REGION Network 2
   RUNG wire#powerrail
      "DB204"(IN0 := "4#配料皮带备妥", IN1 := "干矿提升皮带运行", IN2 :=, IN3 :=, IN4 := "4#配料皮带运行", IN5 :=, OUT6 := "4#配料皮带启动")
      "DB205"(IN0 := "5#配料皮带备妥", IN1 := "干矿提升皮带运行", IN2 :=, IN3 :=, IN4 := "5#配料皮带运行", IN5 :=, OUT6 := "5#配料皮带启动")
      "DB206"(IN0 := "6#配料皮带备妥", IN1 := "干矿提升皮带运行", IN2 :=, IN3 :=, IN4 := "6#配料皮带运行", IN5 :=, OUT6 := "6#配料皮带启动")
   END_RUNG
   // the same network as SCL:
   "DB204"(IN0 := "4#配料皮带备妥", IN1 := "干矿提升皮带运行", IN4 := "4#配料皮带运行", OUT6 := "4#配料皮带启动", ENO => #_w1);   // "给料电机启动块"
   "DB205"(EN := #_w1, IN0 := "5#配料皮带备妥", IN1 := "干矿提升皮带运行", IN4 := "5#配料皮带运行", OUT6 := "5#配料皮带启动", ENO => #_w2);   // "给料电机启动块"
   IF #_w2 THEN
       "DB206"(IN0 := "6#配料皮带备妥", IN1 := "干矿提升皮带运行", IN4 := "6#配料皮带运行", OUT6 := "6#配料皮带启动");   // "给料电机启动块"
   END_IF;
END_REGION

REGION Network 3
   RUNG wire#powerrail
      "DB207"(IN0 := "7#配料皮带备妥", IN1 := "干矿提升皮带运行", IN2 :=, IN3 :=, IN4 := "7#配料皮带运行", IN5 :=, OUT6 := "7#配料皮带启动")
      "DB208"(IN0 := "1#板式给料机备妥", IN1 := "1#板式给料机备妥", IN2 :=, IN3 :=, IN4 := "1#板式给料机运行", IN5 :=, OUT6 := "板式给料机启动")
   END_RUNG
   // the same network as SCL:
   "DB207"(IN0 := "7#配料皮带备妥", IN1 := "干矿提升皮带运行", IN4 := "7#配料皮带运行", OUT6 := "7#配料皮带启动", ENO => #_w1);   // "给料电机启动块"
   IF #_w1 THEN
       "DB208"(IN0 := "1#板式给料机备妥", IN1 := "1#板式给料机备妥", IN4 := "1#板式给料机运行", OUT6 := "板式给料机启动");   // "给料电机启动块"
   END_IF;
END_REGION

REGION Network 4
   RUNG wire#powerrail
      Contact( "DB208".IN3 )
      wire#w1
      I_Contact( "DB208".IN2 )
      Coil( "Q6_7" )
   END_RUNG
   RUNG wire#powerrail
      Contact( "Q6_7" )
   END_RUNG wire#w1
   // the same network as SCL:
   "Q6_7" := ("DB208".IN3 OR "Q6_7") AND NOT "DB208".IN2;
END_REGION
END_FUNCTION

FUNCTION "配料模拟量" : Void   // FC22, LAD
{ S7_Optimized_Access := 'FALSE' }
VERSION : 0.1
BEGIN

REGION Network 1
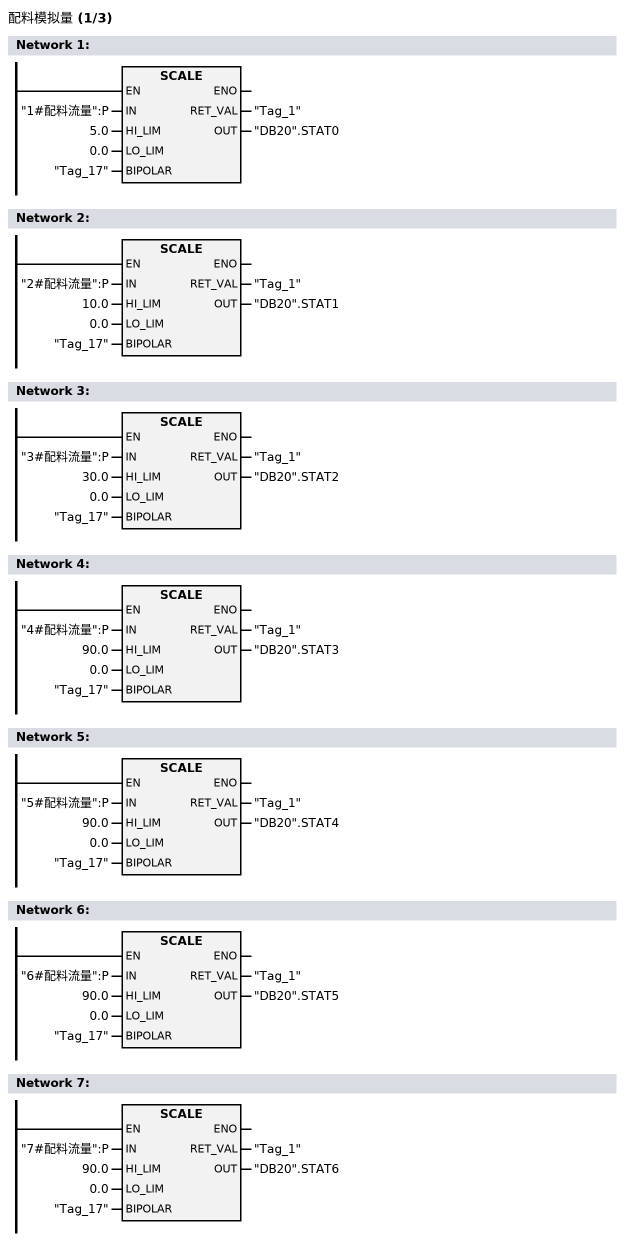
   "Tag_1" := SCALE(IN := "1#配料流量":P, HI_LIM := 5.0, LO_LIM := 0.0, BIPOLAR := "Tag_17", OUT => "DB20".STAT0);
END_REGION

REGION Network 2
   "Tag_1" := SCALE(IN := "2#配料流量":P, HI_LIM := 10.0, LO_LIM := 0.0, BIPOLAR := "Tag_17", OUT => "DB20".STAT1);
END_REGION

REGION Network 3
   "Tag_1" := SCALE(IN := "3#配料流量":P, HI_LIM := 30.0, LO_LIM := 0.0, BIPOLAR := "Tag_17", OUT => "DB20".STAT2);
END_REGION

REGION Network 4
   "Tag_1" := SCALE(IN := "4#配料流量":P, HI_LIM := 90.0, LO_LIM := 0.0, BIPOLAR := "Tag_17", OUT => "DB20".STAT3);
END_REGION

REGION Network 5
   "Tag_1" := SCALE(IN := "5#配料流量":P, HI_LIM := 90.0, LO_LIM := 0.0, BIPOLAR := "Tag_17", OUT => "DB20".STAT4);
END_REGION

REGION Network 6
   "Tag_1" := SCALE(IN := "6#配料流量":P, HI_LIM := 90.0, LO_LIM := 0.0, BIPOLAR := "Tag_17", OUT => "DB20".STAT5);
END_REGION

REGION Network 7
   "Tag_1" := SCALE(IN := "7#配料流量":P, HI_LIM := 90.0, LO_LIM := 0.0, BIPOLAR := "Tag_17", OUT => "DB20".STAT6);
END_REGION

REGION Network 8
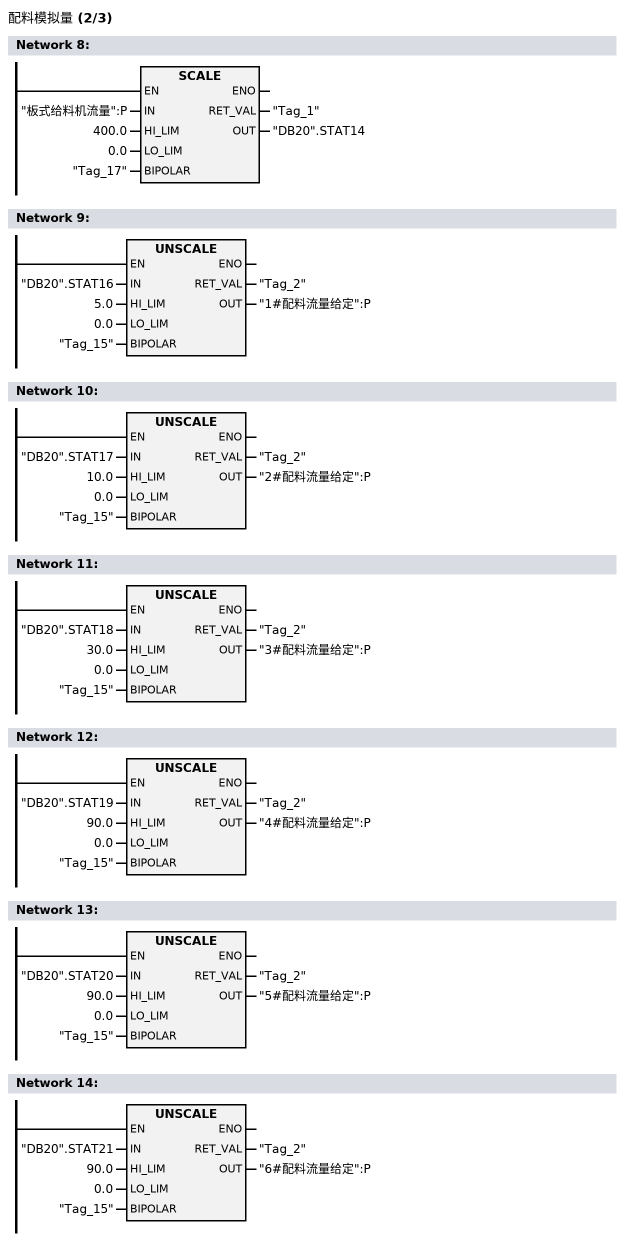
   "Tag_1" := SCALE(IN := "板式给料机流量":P,
                    HI_LIM := 400.0,
                    LO_LIM := 0.0,
                    BIPOLAR := "Tag_17",
                    OUT => "DB20".STAT14);
END_REGION

REGION Network 9
   "Tag_2" := UNSCALE(IN := "DB20".STAT16,
                      HI_LIM := 5.0,
                      LO_LIM := 0.0,
                      BIPOLAR := "Tag_15",
                      OUT => "1#配料流量给定":P);
END_REGION

REGION Network 10
   "Tag_2" := UNSCALE(IN := "DB20".STAT17,
                      HI_LIM := 10.0,
                      LO_LIM := 0.0,
                      BIPOLAR := "Tag_15",
                      OUT => "2#配料流量给定":P);
END_REGION

REGION Network 11
   "Tag_2" := UNSCALE(IN := "DB20".STAT18,
                      HI_LIM := 30.0,
                      LO_LIM := 0.0,
                      BIPOLAR := "Tag_15",
                      OUT => "3#配料流量给定":P);
END_REGION

REGION Network 12
   "Tag_2" := UNSCALE(IN := "DB20".STAT19,
                      HI_LIM := 90.0,
                      LO_LIM := 0.0,
                      BIPOLAR := "Tag_15",
                      OUT => "4#配料流量给定":P);
END_REGION

REGION Network 13
   "Tag_2" := UNSCALE(IN := "DB20".STAT20,
                      HI_LIM := 90.0,
                      LO_LIM := 0.0,
                      BIPOLAR := "Tag_15",
                      OUT => "5#配料流量给定":P);
END_REGION

REGION Network 14
   "Tag_2" := UNSCALE(IN := "DB20".STAT21,
                      HI_LIM := 90.0,
                      LO_LIM := 0.0,
                      BIPOLAR := "Tag_15",
                      OUT => "6#配料流量给定":P);
END_REGION

REGION Network 15
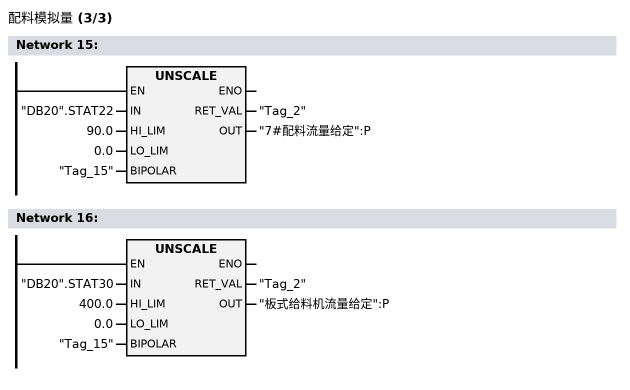
   "Tag_2" := UNSCALE(IN := "DB20".STAT22,
                      HI_LIM := 90.0,
                      LO_LIM := 0.0,
                      BIPOLAR := "Tag_15",
                      OUT => "7#配料流量给定":P);
END_REGION

REGION Network 16
   "Tag_2" := UNSCALE(IN := "DB20".STAT30,
                      HI_LIM := 400.0,
                      LO_LIM := 0.0,
                      BIPOLAR := "Tag_15",
                      OUT => "板式给料机流量给定":P);
END_REGION
END_FUNCTION

FUNCTION "配料累计" : Void   // FC23, LAD
{ S7_Optimized_Access := 'FALSE' }
VERSION : 0.1
   VAR_TEMP   // added for the SCL form of the ladder/FBD networks
      _w1 : Bool;
   END_VAR
BEGIN

REGION Network 1
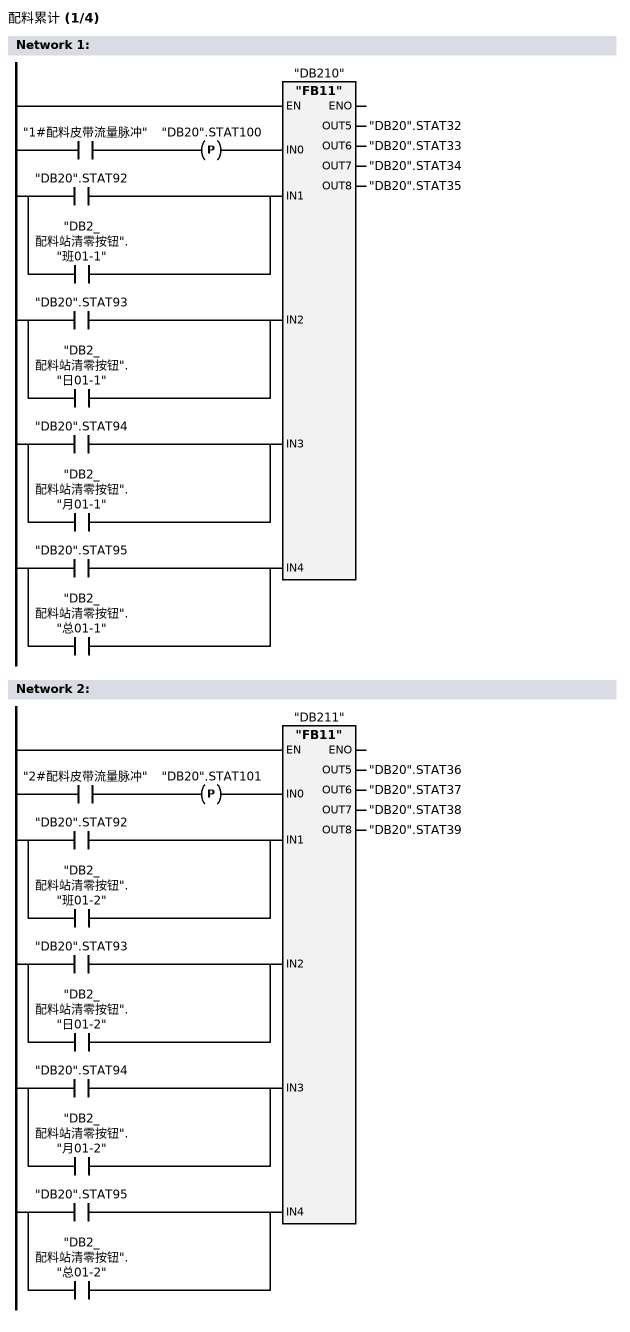
   RUNG wire#powerrail
      "DB210"(IN0 := wire#w1, IN1 := wire#w2, IN2 := wire#w3, IN3 := wire#w4, IN4 := wire#w5, OUT5 => "DB20".STAT32, OUT6 => "DB20".STAT33, OUT7 => "DB20".STAT34, OUT8 => "DB20".STAT35)
   END_RUNG
   RUNG wire#powerrail
      Contact( "1#配料皮带流量脉冲" )
      P_Trig( "DB20".STAT100 )
   END_RUNG wire#w1
   RUNG wire#powerrail
      Contact( "DB20".STAT92 )
   END_RUNG wire#w2
   RUNG wire#powerrail
      Contact( "DB2_配料站清零按钮"."班01-1" )
   END_RUNG wire#w2
   RUNG wire#powerrail
      Contact( "DB20".STAT93 )
   END_RUNG wire#w3
   RUNG wire#powerrail
      Contact( "DB2_配料站清零按钮"."日01-1" )
   END_RUNG wire#w3
   RUNG wire#powerrail
      Contact( "DB20".STAT94 )
   END_RUNG wire#w4
   RUNG wire#powerrail
      Contact( "DB2_配料站清零按钮"."月01-1" )
   END_RUNG wire#w4
   RUNG wire#powerrail
      Contact( "DB20".STAT95 )
   END_RUNG wire#w5
   RUNG wire#powerrail
      Contact( "DB2_配料站清零按钮"."总01-1" )
   END_RUNG wire#w5
   // the same network as SCL:
   #_w1 := "1#配料皮带流量脉冲" AND NOT "DB20".STAT100;   // rising edge
   "DB20".STAT100 := "1#配料皮带流量脉冲";
   "DB210"(IN0 := #_w1,   // "FB11"
           IN1 := "DB20".STAT92 OR "DB2_配料站清零按钮"."班01-1",
           IN2 := "DB20".STAT93 OR "DB2_配料站清零按钮"."日01-1",
           IN3 := "DB20".STAT94 OR "DB2_配料站清零按钮"."月01-1",
           IN4 := "DB20".STAT95 OR "DB2_配料站清零按钮"."总01-1",
           OUT5 => "DB20".STAT32,
           OUT6 => "DB20".STAT33,
           OUT7 => "DB20".STAT34,
           OUT8 => "DB20".STAT35);
END_REGION

REGION Network 2
   RUNG wire#powerrail
      "DB211"(IN0 := wire#w1, IN1 := wire#w2, IN2 := wire#w3, IN3 := wire#w4, IN4 := wire#w5, OUT5 => "DB20".STAT36, OUT6 => "DB20".STAT37, OUT7 => "DB20".STAT38, OUT8 => "DB20".STAT39)
   END_RUNG
   RUNG wire#powerrail
      Contact( "2#配料皮带流量脉冲" )
      P_Trig( "DB20".STAT101 )
   END_RUNG wire#w1
   RUNG wire#powerrail
      Contact( "DB20".STAT92 )
   END_RUNG wire#w2
   RUNG wire#powerrail
      Contact( "DB2_配料站清零按钮"."班01-2" )
   END_RUNG wire#w2
   RUNG wire#powerrail
      Contact( "DB20".STAT93 )
   END_RUNG wire#w3
   RUNG wire#powerrail
      Contact( "DB2_配料站清零按钮"."日01-2" )
   END_RUNG wire#w3
   RUNG wire#powerrail
      Contact( "DB20".STAT94 )
   END_RUNG wire#w4
   RUNG wire#powerrail
      Contact( "DB2_配料站清零按钮"."月01-2" )
   END_RUNG wire#w4
   RUNG wire#powerrail
      Contact( "DB20".STAT95 )
   END_RUNG wire#w5
   RUNG wire#powerrail
      Contact( "DB2_配料站清零按钮"."总01-2" )
   END_RUNG wire#w5
   // the same network as SCL:
   #_w1 := "2#配料皮带流量脉冲" AND NOT "DB20".STAT101;   // rising edge
   "DB20".STAT101 := "2#配料皮带流量脉冲";
   "DB211"(IN0 := #_w1,   // "FB11"
           IN1 := "DB20".STAT92 OR "DB2_配料站清零按钮"."班01-2",
           IN2 := "DB20".STAT93 OR "DB2_配料站清零按钮"."日01-2",
           IN3 := "DB20".STAT94 OR "DB2_配料站清零按钮"."月01-2",
           IN4 := "DB20".STAT95 OR "DB2_配料站清零按钮"."总01-2",
           OUT5 => "DB20".STAT36,
           OUT6 => "DB20".STAT37,
           OUT7 => "DB20".STAT38,
           OUT8 => "DB20".STAT39);
END_REGION

REGION Network 3
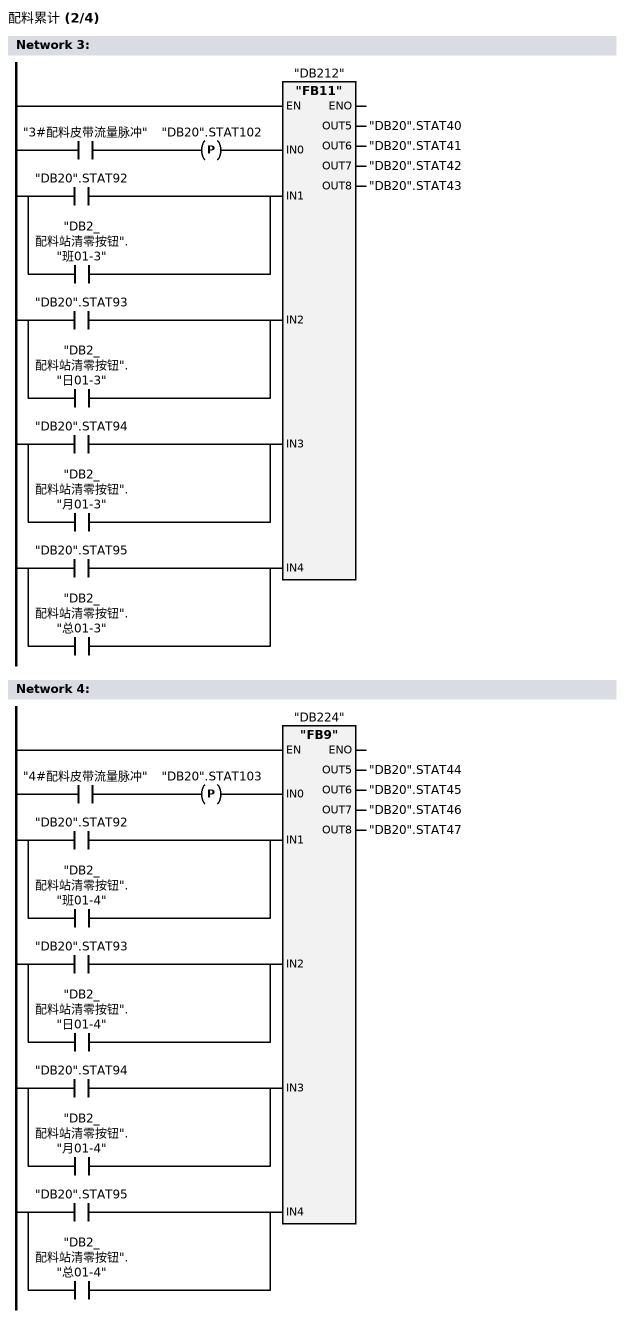
   RUNG wire#powerrail
      "DB212"(IN0 := wire#w1, IN1 := wire#w2, IN2 := wire#w3, IN3 := wire#w4, IN4 := wire#w5, OUT5 => "DB20".STAT40, OUT6 => "DB20".STAT41, OUT7 => "DB20".STAT42, OUT8 => "DB20".STAT43)
   END_RUNG
   RUNG wire#powerrail
      Contact( "3#配料皮带流量脉冲" )
      P_Trig( "DB20".STAT102 )
   END_RUNG wire#w1
   RUNG wire#powerrail
      Contact( "DB20".STAT92 )
   END_RUNG wire#w2
   RUNG wire#powerrail
      Contact( "DB2_配料站清零按钮"."班01-3" )
   END_RUNG wire#w2
   RUNG wire#powerrail
      Contact( "DB20".STAT93 )
   END_RUNG wire#w3
   RUNG wire#powerrail
      Contact( "DB2_配料站清零按钮"."日01-3" )
   END_RUNG wire#w3
   RUNG wire#powerrail
      Contact( "DB20".STAT94 )
   END_RUNG wire#w4
   RUNG wire#powerrail
      Contact( "DB2_配料站清零按钮"."月01-3" )
   END_RUNG wire#w4
   RUNG wire#powerrail
      Contact( "DB20".STAT95 )
   END_RUNG wire#w5
   RUNG wire#powerrail
      Contact( "DB2_配料站清零按钮"."总01-3" )
   END_RUNG wire#w5
   // the same network as SCL:
   #_w1 := "3#配料皮带流量脉冲" AND NOT "DB20".STAT102;   // rising edge
   "DB20".STAT102 := "3#配料皮带流量脉冲";
   "DB212"(IN0 := #_w1,   // "FB11"
           IN1 := "DB20".STAT92 OR "DB2_配料站清零按钮"."班01-3",
           IN2 := "DB20".STAT93 OR "DB2_配料站清零按钮"."日01-3",
           IN3 := "DB20".STAT94 OR "DB2_配料站清零按钮"."月01-3",
           IN4 := "DB20".STAT95 OR "DB2_配料站清零按钮"."总01-3",
           OUT5 => "DB20".STAT40,
           OUT6 => "DB20".STAT41,
           OUT7 => "DB20".STAT42,
           OUT8 => "DB20".STAT43);
END_REGION

REGION Network 4
   RUNG wire#powerrail
      "DB224"(IN0 := wire#w1, IN1 := wire#w2, IN2 := wire#w3, IN3 := wire#w4, IN4 := wire#w5, OUT5 => "DB20".STAT44, OUT6 => "DB20".STAT45, OUT7 => "DB20".STAT46, OUT8 => "DB20".STAT47)
   END_RUNG
   RUNG wire#powerrail
      Contact( "4#配料皮带流量脉冲" )
      P_Trig( "DB20".STAT103 )
   END_RUNG wire#w1
   RUNG wire#powerrail
      Contact( "DB20".STAT92 )
   END_RUNG wire#w2
   RUNG wire#powerrail
      Contact( "DB2_配料站清零按钮"."班01-4" )
   END_RUNG wire#w2
   RUNG wire#powerrail
      Contact( "DB20".STAT93 )
   END_RUNG wire#w3
   RUNG wire#powerrail
      Contact( "DB2_配料站清零按钮"."日01-4" )
   END_RUNG wire#w3
   RUNG wire#powerrail
      Contact( "DB20".STAT94 )
   END_RUNG wire#w4
   RUNG wire#powerrail
      Contact( "DB2_配料站清零按钮"."月01-4" )
   END_RUNG wire#w4
   RUNG wire#powerrail
      Contact( "DB20".STAT95 )
   END_RUNG wire#w5
   RUNG wire#powerrail
      Contact( "DB2_配料站清零按钮"."总01-4" )
   END_RUNG wire#w5
   // the same network as SCL:
   #_w1 := "4#配料皮带流量脉冲" AND NOT "DB20".STAT103;   // rising edge
   "DB20".STAT103 := "4#配料皮带流量脉冲";
   "DB224"(IN0 := #_w1,   // "FB9"
           IN1 := "DB20".STAT92 OR "DB2_配料站清零按钮"."班01-4",
           IN2 := "DB20".STAT93 OR "DB2_配料站清零按钮"."日01-4",
           IN3 := "DB20".STAT94 OR "DB2_配料站清零按钮"."月01-4",
           IN4 := "DB20".STAT95 OR "DB2_配料站清零按钮"."总01-4",
           OUT5 => "DB20".STAT44,
           OUT6 => "DB20".STAT45,
           OUT7 => "DB20".STAT46,
           OUT8 => "DB20".STAT47);
END_REGION

REGION Network 5
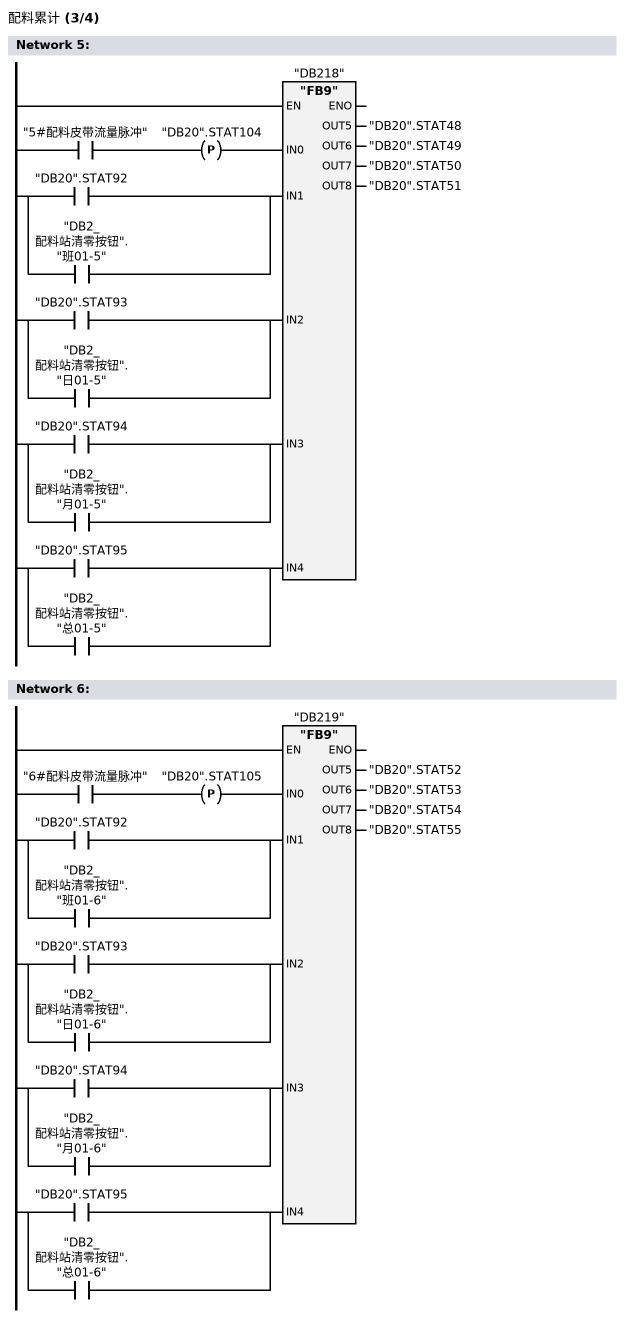
   RUNG wire#powerrail
      "DB218"(IN0 := wire#w1, IN1 := wire#w2, IN2 := wire#w3, IN3 := wire#w4, IN4 := wire#w5, OUT5 => "DB20".STAT48, OUT6 => "DB20".STAT49, OUT7 => "DB20".STAT50, OUT8 => "DB20".STAT51)
   END_RUNG
   RUNG wire#powerrail
      Contact( "5#配料皮带流量脉冲" )
      P_Trig( "DB20".STAT104 )
   END_RUNG wire#w1
   RUNG wire#powerrail
      Contact( "DB20".STAT92 )
   END_RUNG wire#w2
   RUNG wire#powerrail
      Contact( "DB2_配料站清零按钮"."班01-5" )
   END_RUNG wire#w2
   RUNG wire#powerrail
      Contact( "DB20".STAT93 )
   END_RUNG wire#w3
   RUNG wire#powerrail
      Contact( "DB2_配料站清零按钮"."日01-5" )
   END_RUNG wire#w3
   RUNG wire#powerrail
      Contact( "DB20".STAT94 )
   END_RUNG wire#w4
   RUNG wire#powerrail
      Contact( "DB2_配料站清零按钮"."月01-5" )
   END_RUNG wire#w4
   RUNG wire#powerrail
      Contact( "DB20".STAT95 )
   END_RUNG wire#w5
   RUNG wire#powerrail
      Contact( "DB2_配料站清零按钮"."总01-5" )
   END_RUNG wire#w5
   // the same network as SCL:
   #_w1 := "5#配料皮带流量脉冲" AND NOT "DB20".STAT104;   // rising edge
   "DB20".STAT104 := "5#配料皮带流量脉冲";
   "DB218"(IN0 := #_w1,   // "FB9"
           IN1 := "DB20".STAT92 OR "DB2_配料站清零按钮"."班01-5",
           IN2 := "DB20".STAT93 OR "DB2_配料站清零按钮"."日01-5",
           IN3 := "DB20".STAT94 OR "DB2_配料站清零按钮"."月01-5",
           IN4 := "DB20".STAT95 OR "DB2_配料站清零按钮"."总01-5",
           OUT5 => "DB20".STAT48,
           OUT6 => "DB20".STAT49,
           OUT7 => "DB20".STAT50,
           OUT8 => "DB20".STAT51);
END_REGION

REGION Network 6
   RUNG wire#powerrail
      "DB219"(IN0 := wire#w1, IN1 := wire#w2, IN2 := wire#w3, IN3 := wire#w4, IN4 := wire#w5, OUT5 => "DB20".STAT52, OUT6 => "DB20".STAT53, OUT7 => "DB20".STAT54, OUT8 => "DB20".STAT55)
   END_RUNG
   RUNG wire#powerrail
      Contact( "6#配料皮带流量脉冲" )
      P_Trig( "DB20".STAT105 )
   END_RUNG wire#w1
   RUNG wire#powerrail
      Contact( "DB20".STAT92 )
   END_RUNG wire#w2
   RUNG wire#powerrail
      Contact( "DB2_配料站清零按钮"."班01-6" )
   END_RUNG wire#w2
   RUNG wire#powerrail
      Contact( "DB20".STAT93 )
   END_RUNG wire#w3
   RUNG wire#powerrail
      Contact( "DB2_配料站清零按钮"."日01-6" )
   END_RUNG wire#w3
   RUNG wire#powerrail
      Contact( "DB20".STAT94 )
   END_RUNG wire#w4
   RUNG wire#powerrail
      Contact( "DB2_配料站清零按钮"."月01-6" )
   END_RUNG wire#w4
   RUNG wire#powerrail
      Contact( "DB20".STAT95 )
   END_RUNG wire#w5
   RUNG wire#powerrail
      Contact( "DB2_配料站清零按钮"."总01-6" )
   END_RUNG wire#w5
   // the same network as SCL:
   #_w1 := "6#配料皮带流量脉冲" AND NOT "DB20".STAT105;   // rising edge
   "DB20".STAT105 := "6#配料皮带流量脉冲";
   "DB219"(IN0 := #_w1,   // "FB9"
           IN1 := "DB20".STAT92 OR "DB2_配料站清零按钮"."班01-6",
           IN2 := "DB20".STAT93 OR "DB2_配料站清零按钮"."日01-6",
           IN3 := "DB20".STAT94 OR "DB2_配料站清零按钮"."月01-6",
           IN4 := "DB20".STAT95 OR "DB2_配料站清零按钮"."总01-6",
           OUT5 => "DB20".STAT52,
           OUT6 => "DB20".STAT53,
           OUT7 => "DB20".STAT54,
           OUT8 => "DB20".STAT55);
END_REGION

REGION Network 7
